// TIA Portal project "YDSLK_HMI_2023-05-10_08-26_V3_00T" (V15.1)

(* hardware
DEVICE "SIMATIC HMI Station_韩国"  TP1200 Comfort
   slot 0: "SIMATIC HMI Station_韩国"  TP1200 Comfort  6AV2 124-0MC01-0AX0  15.0.0.0
   slot 1: "WinCC flexible RT_1"  TP1200 Comfort  6AV2 124-0MC01-0AX0  15.0.0.0
   slot 5: "SIMATIC HMI Station_韩国..IE_CP_1"  PROFINET Interface  15.0.0.0
      slot 1: "PROFINET Interface_1"  PROFINET Interface
         slot 1: "Port_1"  Port
         slot 2: "Port_2"  Port
   slot 7: "SIMATIC HMI Station_韩国..MPI/DP_CP_1"  MPI/DP Interface  15.0.0.0
DEVICE "DeviceProxy-Station_2"  DeviceProxy-Station
   slot 0: "机架_0"  Rail
   slot 1: "DP"  SIMOTION
   slot 2: "DP/MPI"  SIMOTION
   slot 2: "PLC_proxy_2_PN"  Device Proxy  D425_2_DPPN_V45_S120_V48_CPU:6AU1 425-2AD00-0AA0  V4.5
   slot 4: "PNxIE-NET"  SIMOTION
      slot 1: "端口_1"  Port
   slot 6: "PNxIO"  SIMOTION
      slot 1: "端口_1"  Port
   slot 15: "PNxIE"  SIMOTION
      slot 1: "端口_1"  Port
DEVICE "DeviceProxy-Station_1"  DeviceProxy-Station
   slot 0: "机架_0"  Rail
   slot 1: "DP"  SIMOTION
   slot 2: "DP/MPI"  SIMOTION
   slot 2: "PLC_proxy_1_DP"  Device Proxy  D425_DP_V45_S120_V48_CPU:6AU1 425-2AA00-0AA0  V4.5
   slot 4: "PNxIE-NET"  SIMOTION
      slot 1: "端口_1"  Port
   slot 11: "PNxIE-OP"  SIMOTION
      slot 1: "端口_1"  Port
   slot 15: "PNxIE"  SIMOTION
      slot 1: "端口_1"  Port
DEVICE "SIMATIC HMI Station_中国"  TP1200 Comfort
   slot 0: "SIMATIC HMI Station_中国"  TP1200 Comfort  6AV2 124-0MC01-0AX0  15.1.0.0
   slot 1: "WinCC flexible RT"  TP1200 Comfort  6AV2 124-0MC01-0AX0  15.1.0.0
   slot 5: "SIMATIC HMI Station(2).IE_CP_1"  PROFINET Interface  15.0.1.0
      slot 1: "PROFINET Interface_1"  PROFINET Interface
         slot 1: "Port_1"  Port
         slot 2: "Port_2"  Port
   slot 7: "SIMATIC HMI Station(2).MPI/DP_CP_1"  MPI/DP Interface  15.0.1.0
*)

// ===== PLC "PLC_proxy_2_PN"  Device Proxy =====

// ===== PLC "PLC_proxy_1_DP"  Device Proxy =====

(* ===== HMI "HMI_RT_1" =====

ScreenModuleEditorView "面板_1(2)" 640x480
   Group "Group" at 10,10 size 111x159
*)

(* ===== HMI "WinCC flexible RT_1" =====
system functions are stored by id; their names below are inferred from use
connection "HMI_连接_2": ETHERNET, SIMOTION

HMI tags "默认变量表"
   "ST_FC_Var_g_Position_ZouChe_Zhangli_mid" : LReal = PLC ST_FC_Var.g_Position_ZouChe_Zhangli_mid AT 10-30-00-01-00-1F-84-04-ED-80, 1 s
   "ST_HMI_Var_HMI_r64Axis_ChengXing_PositiveAccel_CunRao" : LReal = PLC ST_HMI_Var.HMI_r64Axis_ChengXing_PositiveAccel_CunRao AT 10-30-00-01-00-21-84-00-3C-40, 1 s
   "ST_Cam5_Data_Var_fi" : LReal = PLC ST_Cam5_Data_Var.fi AT 10-30-00-01-00-17-84-00-05-00, 1 s
   "ST_HMI_Var_HMI_r64QianShen_FenSan_real" : LReal = PLC ST_HMI_Var.HMI_r64QianShen_FenSan_real AT 10-30-00-01-00-21-84-00-6E-C0, 100 ms
   "ST_HMI_Var_HMI_i_Z" : LReal = PLC ST_HMI_Var.HMI_i_Z AT 10-30-00-01-00-21-84-00-43-40, 1 s
   "ST_HMI_Var_HMI_r64_cam_ChengXing_negativeaccelendjerk_tuirao" : LReal = PLC ST_HMI_Var.HMI_r64_cam_ChengXing_negativeaccelendjerk_tuirao AT 10-30-00-01-00-21-84-00-32-00, 1 s
   "ST_HMI_Var_HMI_r64Axis_ZouChe_negativeaccelendjerk_JinChe" : LReal = PLC ST_HMI_Var.HMI_r64Axis_ZouChe_negativeaccelendjerk_JinChe AT 10-30-00-01-00-21-84-00-15-80, 1 s
   "ST_HMI_Var_HMI_bo_INF_Feed_ON_OFF_Status" : Bool = PLC ST_HMI_Var.HMI_bo_INF_Feed_ON_OFF_Status AT 10-01-00-01-00-21-84-00-72-38, 1 s
   "变量_24" : Int, internal
   "ST_HMI_Var_HMI_r64Position_NianSuo" : LReal = PLC ST_HMI_Var.HMI_r64Position_NianSuo AT 10-30-00-01-00-21-84-00-04-C0, 1 s
   "ST_HMI_Var_HMI_r64NianDu_real" : LReal = PLC ST_HMI_Var.HMI_r64NianDu_real AT 10-30-00-01-00-21-84-00-6D-C0, 100 ms
   "ST_HMI_Var_HMI_r64_LuoSha_PositiveAccel_ZhangLi_FangKai" : LReal = PLC ST_HMI_Var.HMI_r64_LuoSha_PositiveAccel_ZhangLi_FangKai AT 10-30-00-01-00-21-84-00-21-40, 1 s
   "ST_HMI_Var_HMI_r64Height_ShaSui_whole" : LReal = PLC ST_HMI_Var.HMI_r64Height_ShaSui_whole AT 10-30-00-01-00-21-84-00-0B-00, 1 s
   "变量_26" : Int, internal
   "ST_HMI_Var_HMI_r64Axis_ZouChe_positiveaccelstartjerk_ChuChe" : LReal = PLC ST_HMI_Var.HMI_r64Axis_ZouChe_positiveaccelstartjerk_ChuChe AT 10-30-00-01-00-21-84-00-13-80, 1 s
   "ST_HMI_Var_HMI_r64Axis_DingZi_PositiveAccel_TuiRao" : LReal = PLC ST_HMI_Var.HMI_r64Axis_DingZi_PositiveAccel_TuiRao AT 10-30-00-01-00-21-84-00-2D-80, 1 s
   "ST_HMI_Var_HMI_r64NianDu_NianSuo" : LReal = PLC ST_HMI_Var.HMI_r64NianDu_NianSuo AT 10-30-00-01-00-21-84-00-04-80, 1 s
   "VBS_maintenanceWarnStatus_1" : UInt, internal
   "ST_HMI_Var_HMI_alpha_JuanRao_2" : LReal = PLC ST_HMI_Var.HMI_alpha_JuanRao_2 AT 10-30-00-01-00-21-84-00-33-40, 1 s
   "ST_HMI_Var_HMI_T_Z_max" : LReal = PLC ST_HMI_Var.HMI_T_Z_max AT 10-30-00-01-00-21-84-00-43-80, 1 s
   "Axis_ZouChe_positioningState_actualPosition" : LReal = PLC Axis_ZouChe.positioningState.actualPosition AT A1-30-00-08-00-0A-00-00-02-23, 1 s   // Actual position of axis
   "ST_HMI_Var_HMI_r64Axis_ChengXing_positiveaccelendjerk_CunRao" : LReal = PLC ST_HMI_Var.HMI_r64Axis_ChengXing_positiveaccelendjerk_CunRao AT 10-30-00-01-00-21-84-00-3C-C0, 1 s
   "VBS_time_all_hour" : LReal, internal
   "ST_HMI_Var_HMI_r64Axis_DingZi_negativeaccelendjerk_TuiRao" : LReal = PLC ST_HMI_Var.HMI_r64Axis_DingZi_negativeaccelendjerk_TuiRao AT 10-30-00-01-00-21-84-00-2E-80, 1 s
   "VBS_j_times_3" : UInt, internal
   "ST_VAR_ZouChe_g_r64Axis_ZouChe_Position_JuanRao_DingZi_Velocity_Set" : LReal = PLC ST_VAR_ZouChe.g_r64Axis_ZouChe_Position_JuanRao_DingZi_Velocity_Set AT 10-30-00-01-00-42-84-00-00-40, 1 s
   "ST_Calculation_Var_g_i16_Calculation_0_3_Select_Status" : Int = PLC ST_Calculation_Var.g_i16_Calculation_0_3_Select_Status AT 10-05-00-01-00-13-84-00-00-80, 1 s
   "ST_HMI_Var_HMI_bo_ShengTou_QiDong" : Bool = PLC ST_HMI_Var.HMI_bo_ShengTou_QiDong AT 10-01-00-01-00-21-84-00-72-20, 1 s
   "ST_HMI_Var_HMI_bo_JiaNian" : Bool = PLC ST_HMI_Var.HMI_bo_JiaNian AT 10-01-00-01-00-21-84-00-6C-00, 1 s
   "ST_HMI_Var_HMI_r64_Hs2_0_delt" : LReal = PLC ST_HMI_Var.HMI_r64_Hs2_0_delt AT 10-30-00-01-00-21-84-00-33-C0, 1 s
   "ST_Main_Var_g_i16_Mode_Selected" : Int = PLC ST_Main_Var.g_i16_Mode_Selected AT 10-05-00-01-00-23-84-00-51-80, 1 s
   "ST_HMI_Var_HMI_r64Axis_DingZi_negativeaccelstartjerk_TuiRao" : LReal = PLC ST_HMI_Var.HMI_r64Axis_DingZi_negativeaccelstartjerk_TuiRao AT 10-30-00-01-00-21-84-00-2E-40, 1 s
   "ST_HMI_Var_HMI_r64Axis_ChengXing_negativeaccelendjerk_TuiRao" : LReal = PLC ST_HMI_Var.HMI_r64Axis_ChengXing_negativeaccelendjerk_TuiRao AT 10-30-00-01-00-21-84-00-27-40, 1 s
   "ST_HMI_Var_HMI_r64Time_JiaNian" : LReal = PLC ST_HMI_Var.HMI_r64Time_JiaNian AT 10-30-00-01-00-21-84-00-03-00, 1 s
   "ST_HMI_Var_HMI_r64Axis_ChengXing_negativeaccelstartjerk_TuiRao" : LReal = PLC ST_HMI_Var.HMI_r64Axis_ChengXing_negativeaccelstartjerk_TuiRao AT 10-30-00-01-00-21-84-00-27-00, 1 s
   "ST_HMI_Var_HMI_r64Axis_DingZi_Velocity_JianShaoZhi" : LReal = PLC ST_HMI_Var.HMI_r64Axis_DingZi_Velocity_JianShaoZhi AT 10-30-00-01-00-21-84-00-2C-80, 1 s
   "VBS_date1" : LReal, internal
   "ST_HMI_Var_HMI_r64Axis_1_ZhangLi_Additive_Torque_TuiRao" : LReal = PLC ST_HMI_Var.HMI_r64Axis_1_ZhangLi_Additive_Torque_TuiRao AT 10-30-00-01-00-21-84-00-2C-40, 1 s
   "ST_HMI_Var_HMI_alpha_JuanRao_1" : LReal = PLC ST_HMI_Var.HMI_alpha_JuanRao_1 AT 10-30-00-01-00-21-84-00-33-00, 1 s
   "ST_HMI_Var_HMI_r64Niandu_all_Current" : LReal = PLC ST_HMI_Var.HMI_r64Niandu_all_Current AT 10-30-00-01-00-21-84-00-01-C0, 1 s
   "ST_HMI_Var_HMI_bo_ZhangLi_CeDing_Start" : Bool = PLC ST_HMI_Var.HMI_bo_ZhangLi_CeDing_Start AT 10-01-00-01-00-21-84-00-72-00, 1 s
   "ST_HMI_Var_HMI_boNianDu_3" : Bool = PLC ST_HMI_Var.HMI_boNianDu_3 AT 10-01-00-01-00-21-84-00-02-C0, 1 s
   "ST_HMI_Var_HMI_r64_ZiDongTingZhi_QianShen_WuNian" : LReal = PLC ST_HMI_Var.HMI_r64_ZiDongTingZhi_QianShen_WuNian AT 10-30-00-01-00-21-84-00-40-40, 1 s
   "ST_VAR_ZhangLi_g_r64Axis_1_ZhangLi_Position_JuanRao_Set" : LReal = PLC ST_VAR_ZhangLi.g_r64Axis_1_ZhangLi_Position_JuanRao_Set AT 10-30-00-01-00-3E-84-00-0A-00, 1 s
   "Axis_ZL_T_FU_positioningState_actualPosition" : LReal = PLC Axis_ZL_T_FU.positioningState.actualPosition AT A1-30-00-08-00-16-00-00-02-23, 1 s   // Actual position of axis
   "ST_MotionTask_cam5_Comb{13}" : LReal = PLC ST_MotionTask_cam5.Comb[13] AT 10-30-00-01-00-26-84-00-0D-80, 1 s
   "变量_11" : UInt, internal
   "ST_Main_Var_g_i16_Automatic_Selected" : Int = PLC ST_Main_Var.g_i16_Automatic_Selected AT 10-05-00-01-00-23-84-00-51-B0, 1 s
   "ST_HMI_Var_HMI_r64Axis_ChengXing_Velocity_TuiRao" : LReal = PLC ST_HMI_Var.HMI_r64Axis_ChengXing_Velocity_TuiRao AT 10-30-00-01-00-21-84-00-26-00, 1 s
   "ST_TO_DZ_FU_Var_HMI_bo_Task_DZ_FU" : Bool = PLC ST_TO_DZ_FU_Var.HMI_bo_Task_DZ_FU AT 10-01-00-01-00-37-84-00-04-D0, 1 s
   "ST_HMI_Var_HMI_r64Axis_ZouChe_Velocity_ZiDongTingZhi" : LReal = PLC ST_HMI_Var.HMI_r64Axis_ZouChe_Velocity_ZiDongTingZhi AT 10-30-00-01-00-21-84-00-41-80, 1 s
   "ST_HMI_Var_sehao" : String[80] = PLC ST_HMI_Var.sehao AT 10-33-00-51-00-21-84-00-68-70, 1 s
   "ST_HMI_Var_HMI_r64Height_ShaSui_Bottom" : LReal = PLC ST_HMI_Var.HMI_r64Height_ShaSui_Bottom AT 10-30-00-01-00-21-84-00-0A-C0, 1 s
   "ST_HMI_Var_HMI_r64Axis_ZouChe_Position_ZiDongTingZhi" : LReal = PLC ST_HMI_Var.HMI_r64Axis_ZouChe_Position_ZiDongTingZhi AT 10-30-00-01-00-21-84-00-41-40, 1 s
   "VBS_maintenanceWarnStatus_7" : UInt, internal
   "ST_HMI_Var_HMI_alpha_TuiRao_5" : LReal = PLC ST_HMI_Var.HMI_alpha_TuiRao_5 AT 10-30-00-01-00-21-84-00-29-80, 1 s
   "ST_HMI_Var_HMI_r64Axis_DingZi_PositiveAccel_ZiDongTingZhi" : LReal = PLC ST_HMI_Var.HMI_r64Axis_DingZi_PositiveAccel_ZiDongTingZhi AT 10-30-00-01-00-21-84-00-42-00, 1 s
   "ST_Cam5_Data_Var_g_vm" : LReal = PLC ST_Cam5_Data_Var.g_vm AT 10-30-00-01-00-17-84-00-00-40, 1 s
   "ST_Cam5_Data_Var_g_ratio" : LReal = PLC ST_Cam5_Data_Var.g_ratio AT 10-30-00-01-00-17-84-00-02-40, 1 s
   "ST_HMI_Var_HMI_cam2_ratio_delt_max" : LReal = PLC ST_HMI_Var.HMI_cam2_ratio_delt_max AT 10-30-00-01-00-21-84-00-30-40, 1 s
   "ST_HMI_Var_HMI_r64Axis_1_ZhangLi_Position_JuanRao_Set_N" : LReal = PLC ST_HMI_Var.HMI_r64Axis_1_ZhangLi_Position_JuanRao_Set_N AT 10-30-00-01-00-21-84-00-39-40, 1 s
   "变量_9" : UInt, internal
   "ST_HMI_Var_HMI_r64_k_ZhangLi_Rate" : LReal = PLC ST_HMI_Var.HMI_r64_k_ZhangLi_Rate AT 10-30-00-01-00-21-84-00-10-C0, 1 s
   "ST_Cam5_Data_Var_sj" : LReal = PLC ST_Cam5_Data_Var.sj AT 10-30-00-01-00-17-84-00-04-00, 1 s
   "ST_HMI_Var_HMI_r64Axis_DingZi_positiveaccelendjerk_JiaNian" : LReal = PLC ST_HMI_Var.HMI_r64Axis_DingZi_positiveaccelendjerk_JiaNian AT 10-30-00-01-00-21-84-00-25-40, 1 s
   "ST_MotionTask_cam5_Comb{2}" : LReal = PLC ST_MotionTask_cam5.Comb[2] AT 10-30-00-01-00-26-84-00-0A-C0, 1 s
   "变量_1" : WString[10], internal
   "ST_Cam5_Data_Var_q" : LReal = PLC ST_Cam5_Data_Var.q AT 10-30-00-01-00-17-84-00-03-40, 1 s
   "ST_HMI_Var_HMI_r64Axis_DingZi_Positiveaccelstartjerk_JiaNian" : LReal = PLC ST_HMI_Var.HMI_r64Axis_DingZi_Positiveaccelstartjerk_JiaNian AT 10-30-00-01-00-21-84-00-25-00, 1 s
   "ST_HMI_Var_HMI_r64Diameter_ShaSui_Max" : LReal = PLC ST_HMI_Var.HMI_r64Diameter_ShaSui_Max AT 10-30-00-01-00-21-84-00-0B-C0, 1 s
   "变量_35" : Bool, internal
   "ST_Main_Var_g_i16_Mode_Enabled" : Int = PLC ST_Main_Var.g_i16_Mode_Enabled AT 10-05-00-01-00-00-82-00-00-50, 1 s
   "VBS_j_times_2" : UInt, internal
   "变量_3" : UInt, internal
   "ST_HMI_Var_HMI_r64Height_ShaGuan_Middle" : LReal = PLC ST_HMI_Var.HMI_r64Height_ShaGuan_Middle AT 10-30-00-01-00-21-84-00-0D-80, 1 s
   "ST_HMI_Var_HMI_cam2_ratio_min" : LReal = PLC ST_HMI_Var.HMI_cam2_ratio_min AT 10-30-00-01-00-21-84-00-2F-40, 1 s
   "Picture" : Int, internal
   "ST_Cam5_Data_Var_s" : LReal = PLC ST_Cam5_Data_Var.s AT 10-30-00-01-00-17-84-00-02-80, 1 s
   "ST_FC_Var_g_g1_n_delt_ratio" : LReal = PLC ST_FC_Var.g_g1_n_delt_ratio AT 10-30-00-01-00-1F-84-04-EB-00, 1 s
   "ST_HMI_Var_HMI_r64Axis_ChengXing_negativeaccelendjerk_CunRao" : LReal = PLC ST_HMI_Var.HMI_r64Axis_ChengXing_negativeaccelendjerk_CunRao AT 10-30-00-01-00-21-84-00-3D-40, 1 s
   "VBS_j_times_6" : UInt, internal
   "ST_HMI_Var_HMI_bo_ChuChe" : Bool = PLC ST_HMI_Var.HMI_bo_ChuChe AT 10-01-00-01-00-21-84-00-6B-D0, 1 s
   "ST_FC_Var_g_f1_n_delt_max" : LReal = PLC ST_FC_Var.g_f1_n_delt_max AT 10-30-00-01-00-1F-84-04-ED-00, 1 s
   "ST_HMI_Var_HMI_r64Time_ChuChe" : LReal = PLC ST_HMI_Var.HMI_r64Time_ChuChe AT 10-30-00-01-00-21-84-00-09-C0, 1 s
   "ST_HMI_Var_HMI_r64QianShen_All_real_ShengTou" : LReal = PLC ST_HMI_Var.HMI_r64QianShen_All_real_ShengTou AT 10-30-00-01-00-21-84-00-71-00, 1 s
   "ST_HMI_Var_HMI_f1_n_delt_new_0" : LReal = PLC ST_HMI_Var.HMI_f1_n_delt_new_0 AT 10-30-00-01-00-21-84-00-39-80, 1 s
   "ST_Cam5_Data_Var_sq1" : LReal = PLC ST_Cam5_Data_Var.sq1 AT 10-30-00-01-00-17-84-00-03-C0, 1 s
   "ST_Main_Var_g_i16_Automatic_Status" : Int = PLC ST_Main_Var.g_i16_Automatic_Status AT 10-05-00-01-00-00-82-00-00-A0, 1 s
   "ST_HMI_Var_HMI_r64Axis_ZouChe_positiveaccelstartjerk_JinChe" : LReal = PLC ST_HMI_Var.HMI_r64Axis_ZouChe_positiveaccelstartjerk_JinChe AT 10-30-00-01-00-21-84-00-14-C0, 1 s
   "ST_HMI_Var_HMI_r64Axis_ChengXing_PositiveAccel_TuiRao" : LReal = PLC ST_HMI_Var.HMI_r64Axis_ChengXing_PositiveAccel_TuiRao AT 10-30-00-01-00-21-84-00-26-40, 1 s
   "ST_HMI_Var_HMI_bo_chuche_select" : Bool = PLC ST_HMI_Var.HMI_bo_chuche_select AT 10-01-00-01-00-21-84-00-08-80, 1 s
   "ST_Main_Var_g_bo_Mode_Enabled_Disable" : Bool = PLC ST_Main_Var.g_bo_Mode_Enabled_Disable AT 10-01-00-01-00-00-82-00-00-59, 1 s
   "ST_HMI_Var_HMI_r64_cam_DingZi_positiveaccel_TuiRao" : LReal = PLC ST_HMI_Var.HMI_r64_cam_DingZi_positiveaccel_TuiRao AT 10-30-00-01-00-21-84-00-2B-40, 1 s
   "ST_HMI_Var_HMI_r64NianDu_3" : LReal = PLC ST_HMI_Var.HMI_r64NianDu_3 AT 10-30-00-01-00-21-84-00-02-80, 1 s
   "变量_29" : Int, internal
   "ST_HMI_Var_HMI_r64_ZiDongTingZhi_QianShen_All" : LReal = PLC ST_HMI_Var.HMI_r64_ZiDongTingZhi_QianShen_All AT 10-30-00-01-00-21-84-00-40-00, 1 s
   "Axis_GunTong_positioningState_actualPosition" : LReal = PLC Axis_GunTong.positioningState.actualPosition AT A1-30-00-08-00-0E-00-00-02-23, 1 s   // Actual position of axis
   "ST_HMI_Var_HMI_r64Time_NianSuo" : LReal = PLC ST_HMI_Var.HMI_r64Time_NianSuo AT 10-30-00-01-00-21-84-00-05-00, 1 s
   "ST_MotionTask_cam5_Comb{1}" : LReal = PLC ST_MotionTask_cam5.Comb[1] AT 10-30-00-01-00-26-84-00-0A-80, 1 s
   "VBS_j_times_7" : UInt, internal
   "ST_HMI_Var_HMI_r64Axis_1_ZhangLi_Position_JuanRao_real" : LReal = PLC ST_HMI_Var.HMI_r64Axis_1_ZhangLi_Position_JuanRao_real AT 10-30-00-01-00-21-84-00-6F-40, 1 s
   "ST_HMI_Var_HMI_r64Axis_DingZi_Velocity_Start_TuiRao" : LReal = PLC ST_HMI_Var.HMI_r64Axis_DingZi_Velocity_Start_TuiRao AT 10-30-00-01-00-21-84-00-2C-C0, 1 s
   "VBS_maintenanceWarnStatus_5" : UInt, internal
   "ST_HMI_Var_HMI_r64_cam_ChengXing_positiveaccelstartjerk_tuirao" : LReal = PLC ST_HMI_Var.HMI_r64_cam_ChengXing_positiveaccelstartjerk_tuirao AT 10-30-00-01-00-21-84-00-31-40, 1 s
   "ST_HMI_Var_HMI_r64Velocity_Jog_TuiRao" : LReal = PLC ST_HMI_Var.HMI_r64Velocity_Jog_TuiRao AT 10-30-00-01-00-21-84-00-1C-00, 1 s
   "ST_HMI_Var_HMI_r64Diameter_ShaGuan_Top" : LReal = PLC ST_HMI_Var.HMI_r64Diameter_ShaGuan_Top AT 10-30-00-01-00-21-84-00-0D-00, 1 s
   "ST_Cam5_Data_Var_g_tz3" : LReal = PLC ST_Cam5_Data_Var.g_tz3 AT 10-30-00-01-00-17-84-00-00-80, 1 s
   "VBS_runningRate" : LReal, internal
   "ST_Cam5_Data_Var_q1" : LReal = PLC ST_Cam5_Data_Var.q1 AT 10-30-00-01-00-17-84-00-03-80, 1 s
   "ST_HMI_Var_chehao" : Int = PLC ST_HMI_Var.chehao AT 10-05-00-01-00-21-84-00-65-D0, 1 s
   "变量_18" : UInt, internal
   "ST_HMI_Var_HMI_r64Axis_1_ZhangLi_PositiveAccel_from_ChengXing_ratio_tuirao" : LReal = PLC ST_HMI_Var.HMI_r64Axis_1_ZhangLi_PositiveAccel_from_ChengXing_ratio_tuirao AT 10-30-00-01-00-21-84-00-2C-00, 1 s
   "ST_Main_Var_g_i16_Start_Position_Status" : Int = PLC ST_Main_Var.g_i16_Start_Position_Status AT 10-05-00-01-00-23-84-00-55-E0, 1 s
   "VBS_maintenanceWarnStatus_4" : UInt, internal
   "ST_Axis_Enable_Test_HMI_bo_Enable_Axis_GunTong" : Bool = PLC ST_Axis_Enable_Test.HMI_bo_Enable_Axis_GunTong AT 10-01-00-01-00-12-84-00-00-B0, 1 s
   "变量_28" : Int, internal
   "ST_HMI_Var_HMI_r64_cam_ChengXing_negativeaccelendjerk_juanrao" : LReal = PLC ST_HMI_Var.HMI_r64_cam_ChengXing_negativeaccelendjerk_juanrao AT 10-30-00-01-00-21-84-00-37-80, 1 s
   "ST_HMI_Var_HMI_r64Velocity_Jog_ZhangLi_Down" : LReal = PLC ST_HMI_Var.HMI_r64Velocity_Jog_ZhangLi_Down AT 10-30-00-01-00-21-84-00-20-40, 1 s
   "ST_HMI_Var_HMI_r64Time_JinChe" : LReal = PLC ST_HMI_Var.HMI_r64Time_JinChe AT 10-30-00-01-00-21-84-00-0A-00, 1 s
   "ST_HMI_Var_HMI_bo_ZhangLi_Down" : Bool = PLC ST_HMI_Var.HMI_bo_ZhangLi_Down AT 10-01-00-01-00-21-84-00-6C-18, 1 s
   "ST_HMI_Var_HMI_f1_n_ZhangLi_Set_PianTiao_0" : LReal = PLC ST_HMI_Var.HMI_f1_n_ZhangLi_Set_PianTiao_0 AT 10-30-00-01-00-21-84-00-3A-40, 1 s
   "ST_HMI_Var_HMI_r64QuanShu_DingZi_TuiRao" : LReal = PLC ST_HMI_Var.HMI_r64QuanShu_DingZi_TuiRao AT 10-30-00-01-00-21-84-00-0F-80, 1 s
   "ST_Cam5_Data_Var_g_ratioT" : LReal = PLC ST_Cam5_Data_Var.g_ratioT AT 10-30-00-01-00-17-84-00-02-00, 1 s
   "ST_HMI_Var_HMI_k_TuiRao" : LReal = PLC ST_HMI_Var.HMI_k_TuiRao AT 10-30-00-01-00-21-84-00-2A-40, 1 s
   "ST_HMI_Var_HMI_r64QianShen_WuNian" : LReal = PLC ST_HMI_Var.HMI_r64QianShen_WuNian AT 10-30-00-01-00-21-84-00-06-40, 1 s
   "ST_Main_Var_g_r64_Time_tuirao" : LReal = PLC ST_Main_Var.g_r64_Time_tuirao AT 10-30-00-01-00-23-84-00-02-00, 1 s
   "ST_MotionTask_cam5_Comb{14}" : LReal = PLC ST_MotionTask_cam5.Comb[14] AT 10-30-00-01-00-26-84-00-0D-C0, 1 s
   "ST_HMI_Var_HMI_bo_ZhangLi_Up" : Bool = PLC ST_HMI_Var.HMI_bo_ZhangLi_Up AT 10-01-00-01-00-21-84-00-6B-F0, 1 s
   "ST_Main_Var_g_bo_Mode_Enabled_Automatic" : Bool = PLC ST_Main_Var.g_bo_Mode_Enabled_Automatic AT 10-01-00-01-00-00-82-00-00-5E, 1 s
   "ST_Main_Var_g_bo_Automatic_Running_Selected" : Bool = PLC ST_Main_Var.g_bo_Automatic_Running_Selected AT 10-01-00-01-00-23-84-00-51-D8, 1 s
   "ST_HMI_Var_HMI_r64ZhiShu_Actual" : LReal = PLC ST_HMI_Var.HMI_r64ZhiShu_Actual AT 10-30-00-01-00-21-84-00-0A-40, 1 s
   "ST_HMI_Var_HMI_r64Axis_1_ZhangLi_Velocity_from_ChengXing_ratio_tuirao" : LReal = PLC ST_HMI_Var.HMI_r64Axis_1_ZhangLi_Velocity_from_ChengXing_ratio_tuirao AT 10-30-00-01-00-21-84-00-2B-C0, 1 s
   "ST_HMI_Var_HMI_r64Axis_ZouChe_positiveaccelendjerk_ChuChe" : LReal = PLC ST_HMI_Var.HMI_r64Axis_ZouChe_positiveaccelendjerk_ChuChe AT 10-30-00-01-00-21-84-00-13-C0, 1 s
   "变量_34" : Bool, internal
   "ST_HMI_Var_HMI_r64_cam_ChengXing_velocity_juanrao" : LReal = PLC ST_HMI_Var.HMI_r64_cam_ChengXing_velocity_juanrao AT 10-30-00-01-00-21-84-00-36-00, 1 s
   "ST_HMI_Var_HMI_r64Axis_DingZi_Velocity_object" : LReal = PLC ST_HMI_Var.HMI_r64Axis_DingZi_Velocity_object AT 10-30-00-01-00-21-84-00-6E-00, 1 s
   "ST_HMI_Var_HMI_r64Velocity_ChuChe" : LReal = PLC ST_HMI_Var.HMI_r64Velocity_ChuChe AT 10-30-00-01-00-21-84-00-09-40, 1 s
   "ST_HMI_Var_HMI_r64_Hs2_D_delt" : LReal = PLC ST_HMI_Var.HMI_r64_Hs2_D_delt AT 10-30-00-01-00-21-84-00-34-00, 1 s
   "ST_HMI_Var_HMI_bo_SongTiao" : Bool = PLC ST_HMI_Var.HMI_bo_SongTiao AT 10-01-00-01-00-21-84-00-6B-D8, 1 s
   "ST_HMI_Var_HMI_r64NianSu_1" : LReal = PLC ST_HMI_Var.HMI_r64NianSu_1 AT 10-30-00-01-00-21-84-00-03-80, 1 s
   "ST_HMI_Var_HMI_r64Axis_ZouChe_negativeaccelstartjerk_ChuChe" : LReal = PLC ST_HMI_Var.HMI_r64Axis_ZouChe_negativeaccelstartjerk_ChuChe AT 10-30-00-01-00-21-84-00-14-00, 1 s
   "ST_Main_Var_g_i16_Disable_Status" : Int = PLC ST_Main_Var.g_i16_Disable_Status AT 10-05-00-01-00-23-84-00-51-90, 1 s
   "VBS_j_times_1" : UInt, internal   // 保养次数显示
   "ST_Main_Var_g_r64_Time_jianian" : LReal = PLC ST_Main_Var.g_r64_Time_jianian AT 10-30-00-01-00-23-84-00-01-C0, 1 s
   "ST_HMI_Var_HMI_r64Axis_ZouChe_Position_real_ShengTou" : LReal = PLC ST_HMI_Var.HMI_r64Axis_ZouChe_Position_real_ShengTou AT 10-30-00-01-00-21-84-00-70-80, 1 s
   "ST_HMI_Var_HMI_r64_cam_ChengXing_positiveaccelendjerk_tuirao" : LReal = PLC ST_HMI_Var.HMI_r64_cam_ChengXing_positiveaccelendjerk_tuirao AT 10-30-00-01-00-21-84-00-31-80, 1 s
   "VBS_time_min" : LReal, internal
   "ST_HMI_Var_HMI_r64_cam_ChengXing_negativeaccel_tuirao" : LReal = PLC ST_HMI_Var.HMI_r64_cam_ChengXing_negativeaccel_tuirao AT 10-30-00-01-00-21-84-00-31-00, 1 s
   "变量_22" : Int, internal
   "ST_HMI_Var_HMI_r64_ZiDongTingZhi_NianSu_SheDing" : LReal = PLC ST_HMI_Var.HMI_r64_ZiDongTingZhi_NianSu_SheDing AT 10-30-00-01-00-21-84-00-41-00, 1 s
   "ST_Axis_Enable_Test_HMI_bo_Enable_Axis_1_ZhangLi" : Bool = PLC ST_Axis_Enable_Test.HMI_bo_Enable_Axis_1_ZhangLi AT 10-01-00-01-00-12-84-00-00-98, 1 s
   "ST_HMI_Var_HMI_X_L_0" : LReal = PLC ST_HMI_Var.HMI_X_L_0 AT 10-30-00-01-00-21-84-00-42-80, 1 s
   "ST_Main_Var_g_u16_N_Cycle_Single" : UInt = PLC ST_Main_Var.g_u16_N_Cycle_Single AT 10-04-00-01-00-23-84-00-00-10, 1 s
   "变量_5" : UInt, internal
   "ST_HMI_Var_HMI_r64_cam_ChengXing_positiveaccel_tuirao" : LReal = PLC ST_HMI_Var.HMI_r64_cam_ChengXing_positiveaccel_tuirao AT 10-30-00-01-00-21-84-00-30-C0, 1 s
   "ST_Main_Var_g_i16_Automatic_Stopping_Selected" : Int = PLC ST_Main_Var.g_i16_Automatic_Stopping_Selected AT 10-05-00-01-00-23-84-00-51-F0, 1 s
   "ST_HMI_Var_HMI_r64Axis_ChengXing_Velocity_CunRao" : LReal = PLC ST_HMI_Var.HMI_r64Axis_ChengXing_Velocity_CunRao AT 10-30-00-01-00-21-84-00-3C-00, 1 s
   "ST_HMI_Var_HMI_r64Velocity_Jog_JuanRao" : LReal = PLC ST_HMI_Var.HMI_r64Velocity_Jog_JuanRao AT 10-30-00-01-00-21-84-00-1C-80, 1 s
   "ST_HMI_Var_HMI_x_TuiRao_0" : LReal = PLC ST_HMI_Var.HMI_x_TuiRao_0 AT 10-30-00-01-00-21-84-00-29-C0, 1 s
   "ST_Main_Var_g_r64Axis_1_ZhangLi_Torque_Limit_Positive" : LReal = PLC ST_Main_Var.g_r64Axis_1_ZhangLi_Torque_Limit_Positive AT 10-30-00-01-00-23-84-00-27-80, 1 s
   "ST_Main_Var_g_r64_Length_One_Minute" : LReal = PLC ST_Main_Var.g_r64_Length_One_Minute AT 10-30-00-01-00-23-84-00-02-80, 1 s
   "ST_HMI_Var_HMI_r64Position_ChuChe" : LReal = PLC ST_HMI_Var.HMI_r64Position_ChuChe AT 10-30-00-01-00-21-84-00-09-00, 1 s
   "VBS_j_times_5" : UInt, internal
   "ST_HMI_Var_HMI_r64Velocity_Jog_SongTiao" : LReal = PLC ST_HMI_Var.HMI_r64Velocity_Jog_SongTiao AT 10-30-00-01-00-21-84-00-1A-C0, 1 s
   "ST_HMI_Var_HMI_r64_Hs2_N_delt" : LReal = PLC ST_HMI_Var.HMI_r64_Hs2_N_delt AT 10-30-00-01-00-21-84-00-34-40, 1 s
   "ST_HMI_Var_HMI_r64_Delt_Position_ZouChe_Cam_1_CunRao" : LReal = PLC ST_HMI_Var.HMI_r64_Delt_Position_ZouChe_Cam_1_CunRao AT 10-30-00-01-00-21-84-00-3D-C0, 1 s
   "ST_HMI_Var_HMI_r64_ZiDongTingZhi_QianShen_FenSan" : LReal = PLC ST_HMI_Var.HMI_r64_ZiDongTingZhi_QianShen_FenSan AT 10-30-00-01-00-21-84-00-40-80, 1 s
   "ST_HMI_Var_HMI_r64_ShuLiang_ShaSui" : LReal = PLC ST_HMI_Var.HMI_r64_ShuLiang_ShaSui AT 10-30-00-01-00-21-84-00-21-C0, 1 s
   "ST_HMI_Var_HMI_r64Velocity_Jog_JiaNian" : LReal = PLC ST_HMI_Var.HMI_r64Velocity_Jog_JiaNian AT 10-30-00-01-00-21-84-00-1B-80, 1 s
   "ST_HMI_Var_HMI_r64Axis_DingZi_Velocity_JuanRao_min" : LReal = PLC ST_HMI_Var.HMI_r64Axis_DingZi_Velocity_JuanRao_min AT 10-30-00-01-00-21-84-00-38-00, 1 s
   "ST_HMI_Var_HMI_bo_ChengXing_Up" : Bool = PLC ST_HMI_Var.HMI_bo_ChengXing_Up AT 10-01-00-01-00-21-84-00-6C-10, 1 s
   "变量_31" : Int, internal
   "ST_HMI_Var_HMI_r64Axis_ZouChe_negativeaccelendjerk_ChuChe" : LReal = PLC ST_HMI_Var.HMI_r64Axis_ZouChe_negativeaccelendjerk_ChuChe AT 10-30-00-01-00-21-84-00-14-40, 1 s
   "ST_HMI_Var_HMI_r64Axis_DingZi_PositiveAccel_JuanRao" : LReal = PLC ST_HMI_Var.HMI_r64Axis_DingZi_PositiveAccel_JuanRao AT 10-30-00-01-00-21-84-00-38-80, 1 s
   "ST_HMI_Var_HMI_x_TuiRao_5" : LReal = PLC ST_HMI_Var.HMI_x_TuiRao_5 AT 10-30-00-01-00-21-84-00-2A-00, 1 s
   "变量_19" : UInt, internal
   "ST_FC_Var_g_g1_n_delt_min" : LReal = PLC ST_FC_Var.g_g1_n_delt_min AT 10-30-00-01-00-1F-84-04-EA-80, 1 s
   "ST_Main_Var_g_r64_Time_chuche" : LReal = PLC ST_Main_Var.g_r64_Time_chuche AT 10-30-00-01-00-23-84-00-01-80, 1 s
   "ST_HMI_Var_HMI_scalevalue_Cam_3" : LReal = PLC ST_HMI_Var.HMI_scalevalue_Cam_3 AT 10-30-00-01-00-21-84-00-2A-C0, 1 s
   "ST_HMI_Var_HMI_bo_JinChe" : Bool = PLC ST_HMI_Var.HMI_bo_JinChe AT 10-01-00-01-00-21-84-00-6B-F8, 1 s
   "ST_HMI_Var_HMI_r64_cam_ChengXing_positiveaccelendjerk_juanrao" : LReal = PLC ST_HMI_Var.HMI_r64_cam_ChengXing_positiveaccelendjerk_juanrao AT 10-30-00-01-00-21-84-00-37-00, 1 s
   "ST_FC_Var_g_g1_n_piantiao_min" : LReal = PLC ST_FC_Var.g_g1_n_piantiao_min AT 10-30-00-01-00-1F-84-04-E9-40, 1 s
   "Cam_5_accessState" : DInt = PLC Cam_5.accessState AT A1-07-00-04-00-1E-00-00-00-45, 1 s   // Access data of the cam
   "变量_12" : UInt, internal
   "ST_HMI_Var_HMI_r64_LuoSha_Velocity_ZhangLi_FangKai" : LReal = PLC ST_HMI_Var.HMI_r64_LuoSha_Velocity_ZhangLi_FangKai AT 10-30-00-01-00-21-84-00-21-00, 1 s
   "ST_Axis_Enable_Test_HMI_bo_Enable_Axis_DingZi" : Bool = PLC ST_Axis_Enable_Test.HMI_bo_Enable_Axis_DingZi AT 10-01-00-01-00-12-84-00-00-B8, 1 s
   "ST_HMI_Var_pihao" : String[80] = PLC ST_HMI_Var.pihao AT 10-33-00-51-00-21-84-00-65-E0, 1 s
   "ST_HMI_Var_HMI_r64Axis_DingZi_negativeaccelstartjerk_JiaNian" : LReal = PLC ST_HMI_Var.HMI_r64Axis_DingZi_negativeaccelstartjerk_JiaNian AT 10-30-00-01-00-21-84-00-25-80, 1 s
   "ST_HMI_Var_HMI_r64QianShen_First" : LReal = PLC ST_HMI_Var.HMI_r64QianShen_First AT 10-30-00-01-00-21-84-00-07-40, 1 s
   "ST_HMI_Var_HMI_r64Axis_ZouChe_Position_object" : LReal = PLC ST_HMI_Var.HMI_r64Axis_ZouChe_Position_object AT 10-30-00-01-00-21-84-00-6D-00, 1 s
   "ST_HMI_Var_HMI_r64AccVelocity_Jog_JinChe" : LReal = PLC ST_HMI_Var.HMI_r64AccVelocity_Jog_JinChe AT 10-30-00-01-00-21-84-00-1A-80, 1 s
   "ST_HMI_Var_HMI_r64Axis_1_ZhangLi_Position_JuanRao_Set_0" : LReal = PLC ST_HMI_Var.HMI_r64Axis_1_ZhangLi_Position_JuanRao_Set_0 AT 10-30-00-01-00-21-84-00-38-C0, 1 s
   "ST_HMI_Var_HMI_bo_ShengTou_TingZhi" : Bool = PLC ST_HMI_Var.HMI_bo_ShengTou_TingZhi AT 10-01-00-01-00-21-84-00-72-28, 1 s
   "ST_Axis_Enable_Test_HMI_bo_Enable_Axis_ChengXing" : Bool = PLC ST_Axis_Enable_Test.HMI_bo_Enable_Axis_ChengXing AT 10-01-00-01-00-12-84-00-00-C0, 1 s
   "ST_HMI_Var_HMI_r64Velocity_Jog_Chuche" : LReal = PLC ST_HMI_Var.HMI_r64Velocity_Jog_Chuche AT 10-30-00-01-00-21-84-00-19-C0, 1 s
   "ST_HMI_Var_HMI_r64Axis_ZouChe_PositiveAccel_ZiDongTingZhi" : LReal = PLC ST_HMI_Var.HMI_r64Axis_ZouChe_PositiveAccel_ZiDongTingZhi AT 10-30-00-01-00-21-84-00-41-C0, 1 s
   "ST_HMI_Var_HMI_bo_ChengXing_Down" : Bool = PLC ST_HMI_Var.HMI_bo_ChengXing_Down AT 10-01-00-01-00-21-84-00-6B-E8, 1 s
   "ST_Main_Var_g_u16_PiShu_Whole" : UInt = PLC ST_Main_Var.g_u16_PiShu_Whole AT 10-04-00-01-00-23-84-00-00-60, 1 s
   "ST_Main_Var_Axis_ChengXing_Mode_Select" : Int = PLC ST_Main_Var.Axis_ChengXing_Mode_Select AT 10-05-00-01-00-23-84-00-57-E0, 1 s
   "ST_HMI_Var_HMI_r64StartPosition_Axis_ZouChe" : LReal = PLC ST_HMI_Var.HMI_r64StartPosition_Axis_ZouChe AT 10-30-00-01-00-21-84-00-17-40, 1 s
   "Axis_DingZi_motionStateData_commandVelocity" : LReal = PLC Axis_DingZi.motionStateData.commandVelocity AT A1-30-00-08-00-0F-00-00-00-6A, 1 s   // Set velocity of the axis
   "user_name" : WString[10], internal
   "VBS_time_year" : LReal, internal
   "ST_HMI_Var_HMI_r64Velocity_JinChe" : LReal = PLC ST_HMI_Var.HMI_r64Velocity_JinChe AT 10-30-00-01-00-21-84-00-09-80, 1 s
   "ST_HMI_Var_HMI_r64QianShen_All_real" : LReal = PLC ST_HMI_Var.HMI_r64QianShen_All_real AT 10-30-00-01-00-21-84-00-6E-80, 100 ms
   "ST_Axis_Enable_Test_HMI_bo_Enable_Axis_LuoLa" : Bool = PLC ST_Axis_Enable_Test.HMI_bo_Enable_Axis_LuoLa AT 10-01-00-01-00-12-84-00-00-A8, 1 s
   "变量_7" : UInt, internal
   "ST_FC_Var_g_g1_n_delt_max" : LReal = PLC ST_FC_Var.g_g1_n_delt_max AT 10-30-00-01-00-1F-84-04-EA-C0, 1 s
   "ST_HMI_Var_HMI_gam_ZhangLi_Set_PianTiao_0" : LReal = PLC ST_HMI_Var.HMI_gam_ZhangLi_Set_PianTiao_0 AT 10-30-00-01-00-21-84-00-3A-80, 1 s
   "ST_HMI_Var_HMI_r64_cam_DingZi_velocity_TuiRao" : LReal = PLC ST_HMI_Var.HMI_r64_cam_DingZi_velocity_TuiRao AT 10-30-00-01-00-21-84-00-2B-00, 1 s
   "ST_HMI_Var_HMI_r64Axis_ChengXing_negativeaccelstartjerk_CunRao" : LReal = PLC ST_HMI_Var.HMI_r64Axis_ChengXing_negativeaccelstartjerk_CunRao AT 10-30-00-01-00-21-84-00-3D-00, 1 s
   "ST_HMI_Var_HMI_r64_cam_ChengXing_negativeaccel_juanrao" : LReal = PLC ST_HMI_Var.HMI_r64_cam_ChengXing_negativeaccel_juanrao AT 10-30-00-01-00-21-84-00-36-80, 1 s
   "ST_Main_Var_g_r64_Time_Once" : LReal = PLC ST_Main_Var.g_r64_Time_Once AT 10-30-00-01-00-23-84-00-01-40, 1 s
   "VBS_j_times_4" : UInt, internal
   "ST_HMI_Var_HMI_n_Change_TuiRao" : Int = PLC ST_HMI_Var.HMI_n_Change_TuiRao AT 10-05-00-01-00-21-84-00-2A-80, 1 s
   "ST_HMI_Var_HMI_r64QianShen_finalArea" : LReal = PLC ST_HMI_Var.HMI_r64QianShen_finalArea AT 10-30-00-01-00-21-84-00-08-00, 1 s
   "ST_HMI_Var_HMI_r64Axis_DingZi_positiveaccelendjerk_TuiRao" : LReal = PLC ST_HMI_Var.HMI_r64Axis_DingZi_positiveaccelendjerk_TuiRao AT 10-30-00-01-00-21-84-00-2E-00, 1 s
   "ST_Main_Var_g_r64Axis_DingZi_PositiveAccel_CunRao" : LReal = PLC ST_Main_Var.g_r64Axis_DingZi_PositiveAccel_CunRao AT 10-30-00-01-00-23-84-00-33-00, 1 s
   "ST_MotionTask_cam5_Comb" : Array [0..15] of LReal = PLC ST_MotionTask_cam5.Comb AT 10-30-00-10-00-26-84-00-0A-80, 1 s
   "ST_HMI_Var_HMI_r64Height_ShaSui_Top_MaxD" : LReal = PLC ST_HMI_Var.HMI_r64Height_ShaSui_Top_MaxD AT 10-30-00-01-00-21-84-00-0B-80, 1 s
   "VBS_maintenanceWarnStatus_6" : UInt, internal
   "ST_HMI_Var_HMI_r64Height_ShaGuan_Top" : LReal = PLC ST_HMI_Var.HMI_r64Height_ShaGuan_Top AT 10-30-00-01-00-21-84-00-0D-C0, 1 s
   "ST_Axis_Enable_Test_HMI_bo_Enable_Axis_ZouChe" : Bool = PLC ST_Axis_Enable_Test.HMI_bo_Enable_Axis_ZouChe AT 10-01-00-01-00-12-84-00-00-90, 1 s
   "ST_HMI_Var_HMI_bo_TuiRao" : Bool = PLC ST_HMI_Var.HMI_bo_TuiRao AT 10-01-00-01-00-21-84-00-6B-E0, 1 s
   "ST_Axis_Enable_Test_HMI_bo_Enable_Infeed" : Bool = PLC ST_Axis_Enable_Test.HMI_bo_Enable_Infeed AT 10-01-00-01-00-12-84-00-00-88, 1 s
   "ST_FC_Var_g_f1_n_delt_min" : LReal = PLC ST_FC_Var.g_f1_n_delt_min AT 10-30-00-01-00-1F-84-04-EC-C0, 1 s
   "ST_HMI_Var_HMI_bo_cam2_ratio_delt_switch" : Bool = PLC ST_HMI_Var.HMI_bo_cam2_ratio_delt_switch AT 10-01-00-01-00-21-84-00-2E-C0, 1 s
   "ST_HMI_Var_HMI_r64QianShen_FenSan" : LReal = PLC ST_HMI_Var.HMI_r64QianShen_FenSan AT 10-30-00-01-00-21-84-00-07-00, 1 s
   "Axis_LuoLa_positioningState_actualPosition" : LReal = PLC Axis_LuoLa.positioningState.actualPosition AT A1-30-00-08-00-11-00-00-02-23, 1 s   // Actual position of axis
   "ST_Main_Var_g_i16_Manual_Status" : Int = PLC ST_Main_Var.g_i16_Manual_Status AT 10-05-00-01-00-23-84-00-51-A0, 1 s
   "ST_Axis_Enable_Test_HMI_bo_Enable_Axis_Enable_Test" : Bool = PLC ST_Axis_Enable_Test.HMI_bo_Enable_Axis_Enable_Test AT 10-01-00-01-00-12-84-00-00-80, 1 s
   "变量_6" : UInt, internal
   "ST_HMI_Var_HMI_boAlarm_NianDu_Time" : Bool = PLC ST_HMI_Var.HMI_boAlarm_NianDu_Time AT 10-01-00-01-00-21-84-00-03-40, 1 s
   "ST_HMI_Var_HMI_g1_n_ZhangLi_Set_PianTiao_0" : LReal = PLC ST_HMI_Var.HMI_g1_n_ZhangLi_Set_PianTiao_0 AT 10-30-00-01-00-21-84-00-3A-00, 1 s
   "ST_HMI_Var_HMI_r64ZhiShu_ChengSha" : LReal = PLC ST_HMI_Var.HMI_r64ZhiShu_ChengSha AT 10-30-00-01-00-21-84-00-08-C0, 1 s
   "VBS_maintenanceWarnStatus_2" : UInt, internal
   "VBS_time_sec" : LReal, internal
   "ST_MotionTask_cam5_Comb{16}" : LReal = PLC ST_MotionTask_cam5.Comb[16] AT 10-30-00-01-00-26-84-00-0E-40, 1 s
   "ST_HMI_Var_HMI_r64PositiveAccel_ZouChe_JinChe" : LReal = PLC ST_HMI_Var.HMI_r64PositiveAccel_ZouChe_JinChe AT 10-30-00-01-00-21-84-00-14-80, 1 s
   "VBS_alwaysFalse" : Bool, internal
   "ST_Main_Var_g_r64_Time_juanrao" : LReal = PLC ST_Main_Var.g_r64_Time_juanrao AT 10-30-00-01-00-23-84-00-02-40, 1 s
   "ST_Cam5_Data_Var_vm" : LReal = PLC ST_Cam5_Data_Var.vm AT 10-30-00-01-00-17-84-00-02-C0, 1 s
   "ST_HMI_Var_HMI_r64Velocity_NianSuo" : LReal = PLC ST_HMI_Var.HMI_r64Velocity_NianSuo AT 10-30-00-01-00-21-84-00-05-40, 1 s
   "VBS_maintenanceWarnStatus_3" : UInt, internal
   "ST_HMI_Var_HMI_r64NianDu_real_ShengTou" : LReal = PLC ST_HMI_Var.HMI_r64NianDu_real_ShengTou AT 10-30-00-01-00-21-84-00-70-C0, 1 s
   "ST_HMI_Var_HMI_GAM_max" : LReal = PLC ST_HMI_Var.HMI_GAM_max AT 10-30-00-01-00-21-84-00-43-00, 1 s
   "ST_HMI_Var_HMI_r64ZhiShu_CuSha" : LReal = PLC ST_HMI_Var.HMI_r64ZhiShu_CuSha AT 10-30-00-01-00-21-84-00-08-40, 1 s
   "VBS_maintenanceWarnStatus_index" : UInt, internal
   "ST_HMI_Var_HMI_r64Velocity_DingZi_TuiRao" : LReal = PLC ST_HMI_Var.HMI_r64Velocity_DingZi_TuiRao AT 10-30-00-01-00-21-84-00-0F-C0, 1 s
   "ST_HMI_Var_HMI_r64Axis_DingZi_PositiveAccel_JiaNian" : LReal = PLC ST_HMI_Var.HMI_r64Axis_DingZi_PositiveAccel_JiaNian AT 10-30-00-01-00-21-84-00-24-80, 1 s
   "ST_Calculation_Var_HMI_bo_Calculation_0_Start" : Bool = PLC ST_Calculation_Var.HMI_bo_Calculation_0_Start AT 10-01-00-01-00-13-84-07-FA-40, 1 s
   "变量_27" : Int, internal
   "ST_HMI_Var_HMI_r64Diameter_ShaGuan_Middle" : LReal = PLC ST_HMI_Var.HMI_r64Diameter_ShaGuan_Middle AT 10-30-00-01-00-21-84-00-0C-C0, 1 s
   "ST_HMI_Var_HMI_r64Velocity_Jog_ChengXing_Down" : LReal = PLC ST_HMI_Var.HMI_r64Velocity_Jog_ChengXing_Down AT 10-30-00-01-00-21-84-00-1D-80, 1 s
   "ST_HMI_Var_HMI_r64NianSu_2" : LReal = PLC ST_HMI_Var.HMI_r64NianSu_2 AT 10-30-00-01-00-21-84-00-03-C0, 1 s
   "ST_HMI_Var_HMI_r64Height_ShaSui_Top" : LReal = PLC ST_HMI_Var.HMI_r64Height_ShaSui_Top AT 10-30-00-01-00-21-84-00-0B-40, 1 s
   "ST_Main_Var_g_bo_Automatic_Status_Mergestop" : Bool = PLC ST_Main_Var.g_bo_Automatic_Status_Mergestop AT 10-01-00-01-00-00-82-00-00-A9, 1 s